FUNCTION_BLOCK "DRIVER_4C"   // FB249, SCL
TITLE = DRIVER_4C
{ S7_Optimized_Access := 'FALSE' }
AUTHOR : hugo
FAMILY : AUTOMAT
NAME : DRIVER4C
VERSION : 1.0
// driver_4C is a multi purpose driver.
// a rising edge on in switches from S0 state S1 and the next edge to state S2 and so on.
// in state S0 all outputs Q are FALSE.
// The stet of the Outputs in any state S? is configurable with setup variables.
// The variables S1..S5 define the states, while the sequence is terminated when a state Variable S? = 0.
// The lower bits 0..3 of the state vars S? are corresponding to the Outputs Q0..Q3
   VAR_INPUT
      IN : Bool;
      RST : Bool;
      Timeout : Time;
      SX : Array[1..7] of Byte;
   END_VAR
   VAR_OUTPUT
      SN : Int;
      Q0 : Bool;
      Q1 : Bool;
      Q2 : Bool;
      Q3 : Bool;
   END_VAR
   VAR
      off : TON;
      edge : Bool;
   END_VAR
   VAR_TEMP
      tSX : Byte;
      _SX AT tSX : Array[0..7] of Bool;
   END_VAR
   // SX[1] := B#16#01;
   // SX[2] := B#16#03;
   // SX[3] := B#16#07;
   // SX[4] := B#16#0F;
BEGIN


   IF #RST OR #off.Q THEN
       #SN := 0;
   ELSIF #IN AND NOT #edge THEN
       #SN := #SN + 1;
       IF #SN > 7 OR #SX[#SN] = 0 THEN #SN := 0; END_IF;
   END_IF;
   #edge := #IN;
   IF #SN > 0 THEN
       #tSX := #SX[#SN];  //so und nicht anders
       #Q0 := #_SX[0];
       #Q1 := #_SX[1];
       #Q2 := #_SX[2];
       #Q3 := #_SX[3];
   ELSE
       #Q0 := FALSE;
       #Q1 := FALSE;
       #Q2 := FALSE;
       #Q3 := FALSE;
   END_IF;

   (* maximaum timeout *)
   IF #Timeout > t#0s THEN #off(IN := #SN > 0, PT := #Timeout); END_IF;


   (* revision history
   hm  23. mar. 2009   rev 1.0
       original version

   *)
END_FUNCTION_BLOCK

FUNCTION "T_PLC_MS" : DWord   // FC64, SCL
TITLE = T_PLC_MS
{ S7_Optimized_Access := 'FALSE' }
AUTHOR : hugo
FAMILY : MEASURE
NAME : T_PLC_MS
VERSION : 1.2
// T_PLC_MS reads the internal PLC timer and return the time, it has the advantage to be able to set a debug mode 
// and speed up the counter to test the plc timer overrun which occurs every 50 days respectively 25 days at siemens S7
// this routine also allows to correct the behavior of s7 where the internal plc counter will not count all 32 bits.
// 
// uses: STIME [FB64],IDB_STIME [DB64]
BEGIN


   "IDB_STIME"(); 
   #T_PLC_MS := "IDB_STIME".tx; 
   (* hier muss die korrektur für step7 stattfinden
   plctime muss den vollen wertebereich von time ausnutzen:
   wenn bei step7 time -24tage bis plus 24 tage ist dann muss der timer auch beim überlauf auf -24tage springen 
   und auf keinen fall auf 0 !!!!
   für siemens muss ein weiterer fb im main eingebunden werden der sicherstellt das alle 32 bits durchgezählt werden.
   es kann nur ein fb sein den er muss sich das oberste (32te) bit merken.
   oder etwa spring s7 bei überlauf auf -24 tage????? dann wäre keine korrektur nötig.
   *)
   IF "debug" THEN
       #T_PLC_MS := DINT_TO_DWORD((DWORD_TO_DINT(SHL(IN:=#T_PLC_MS,N:="N") OR SHL(IN:=DWORD#1,N:="N"))-1) + DWORD_TO_DINT("offset_1"));
   END_IF;


   (* revision history
   hm  14.9.2007   rev 1.0
       original version

   hm  12. nov 2007    rev 1.1
       added temporaray variable tx because some compilers could not handle time() as an argument

   hm  16. nov. 2008   rev 1.2
       initialized constants with 0 for compatibility reasons
   *)
END_FUNCTION

FUNCTION "T_PLC_US" : DWord   // FC65, SCL
TITLE = T_PLC_US
{ S7_Optimized_Access := 'FALSE' }
AUTHOR : hugo
FAMILY : MEASURE
NAME : T_PLC_US
VERSION : 1.2
// T_PLC_US reads the internal PLC timer and return the time, it has the advantage to be able to set a debug mode 
// and speed up the counter to test the plc timer overrun which occurs every 50 days respectively 25 days at siemens S7
// this routine also allows to correct the behavior of s7 where the internal plc counter will not count all 32 bits.
// 
// uses: STIME [FB64],IDB_STIME [DB64]
BEGIN


   "IDB_STIME"(); 
   #T_PLC_US := DINT_TO_DWORD(DWORD_TO_DINT("IDB_STIME".tx) * 1000); 
   (* hier muss die korrektur für step7 stattfinden
   plctime muss den vollen wertebereich von time ausnutzen:
   wenn bei step7 time -24tage bis plus 24 tage ist dann muss der timer auch beim überlauf auf -24tage springen 
   und auf keinen fall auf 0 !!!!
   für siemens muss ein weiterer fb im main eingebunden werden der sicherstellt das alle 32 bits durchgezählt werden.
   es kann nur ein fb sein den er muss sich das oberste (32te) bit merken.
   oder etwa spring s7 bei überlauf auf -24 tage????? dann wäre keine korrektur nötig.
   *)
   IF "debug" THEN
       #T_PLC_US := DINT_TO_DWORD((DWORD_TO_DINT(SHL(IN:=#T_PLC_US,N:="N") OR SHL(IN:=DWORD#1,N:="N"))-1) + DWORD_TO_DINT("offset_1"));
   END_IF;


   (* revision history
   hm  14.9.2007   rev 1.0
       original version

   hm  12. nov 2007    rev 1.1
       added temporaray variable tx because some compilers could not handle time() as an argument

   hm  16. nov. 2008   rev 1.2
       initialized constants with 0 for compatibility reasons

   *)
END_FUNCTION

FUNCTION "INC" : Int   // FC90, SCL
TITLE = INC
{ S7_Optimized_Access := 'FALSE' }
AUTHOR : hugo
FAMILY : MATH
NAME : INC
VERSION : 1.1
// This is a increment function which increments the input X by the value D and compares the result with M.
// if the output exceeds M it will continue to count from 0 again.
   VAR_INPUT
      X : Int;
      D : Int;
      "M" : Int;
   END_VAR
BEGIN


     #INC := (#X + #D + #"M" + 1) MOD (#"M" + 1);

   (* revision history
   hm  7. feb 2007   REV 1.0
     original version

   hm  15. jan 2008  rev 1.1
     allow for neagtive increment

   *)
END_FUNCTION

FUNCTION "MULTIME" : Time   // FC203, SCL
TITLE = MULTIME
{ S7_Optimized_Access := 'FALSE' }
AUTHOR : hugo
FAMILY : TIDT
NAME : MULTIME
VERSION : 1.1
// multiplies a time by a real number and returns a time
   VAR_INPUT
      t : Time;
      "M" : Real;
   END_VAR
BEGIN


     #MULTIME := T_CONV(REAL_TO_DINT(DINT_TO_REAL(T_CONV(#t))*#"M"));

   (* revision history
   hm      2. oct 2006 rev 1.0
       original version

   hm      14. mar 2008    rev 1.1
       rounded the result after the last digit

   *)
END_FUNCTION

FUNCTION "MANUAL" : Bool   // FC409, SCL
TITLE = MANUAL
{ S7_Optimized_Access := 'FALSE' }
AUTHOR : hugo
FAMILY : AUTOMAT
NAME : MANUAL
VERSION : 1.0
// MANUAL is a manual override for digital signals.
// when on and off = FALSE, the output follows IN.
// ON = TRUE forces the output high, and OFF = TRUE forces the output low.
   VAR_INPUT
      IN : Bool;
      ON : Bool;
      OFF : Bool;
   END_VAR
BEGIN


   #MANUAL := NOT #OFF AND (#IN OR #ON);


   (* revision history
   hm  21. nov 2008    rev 1.0
       original version


   *)
END_FUNCTION

// ===== PLC "Engineering control"  Unspecific CPU S7 300 =====

VAR_GLOBAL CONSTANT   // PLC tag table "STEP7 classic symbols"
   "debug" : Bool := FALSE;
   "N" : Int := 0;
   "offset" : Int := 0;
   "offset_1" : DWord := 0;
END_VAR

TYPE "REAL2"
VERSION : 0.0
   STRUCT
      R1 : Real;
      RX : Real;
   END_STRUCT;
END_TYPE

DATA_BLOCK "IDB_STIME"   // DB64
{ S7_Optimized_Access := 'FALSE' }
AUTHOR : dalbi
FAMILY : MEASURE
VERSION : 0.0
// stored: InstanceOfName STIME
"STIME"
BEGIN
END_DATA_BLOCK

FUNCTION_BLOCK "CLK_PRG"   // FB52, SCL
TITLE = CLK_PRG
{ S7_Optimized_Access := 'FALSE' }
AUTHOR : hugo
FAMILY : GENERAT
NAME : CLK_PRG
VERSION : 1.3
// clk_prg uses the internal sps time to generate a clock with programmable period time.
// the period time is defined for 10ms .. 65s
// the first cycle after start is a clk pulse and then depending on the programmed period time a delay.
// every pulse is only valid for one cycle.
// the accuracy of clk_prg is depending on the accuracy of the system clock.
// 
// uses: T_PLC_MS [FC64]
//       STIME [FB64],IDB_STIME [DB64]
   VAR_INPUT
      PT : Time := T#10MS;
   END_VAR
   VAR_OUTPUT
      Q : Bool;
   END_VAR
   VAR
      init : Bool;
      last : Time;
      tx : Time;
   END_VAR
   VAR_TEMP
      TOP_SI : Struct
         EV_CLASS : Byte;
         EV_NUM : Byte;
         PRIORITY : Byte;
         NUM : Byte;
         TYP2_3 : Byte;
         TYP1 : Byte;
         ZI1 : Word;
         ZI2_3 : DWord;
      END_STRUCT;
      START_UP_SI : Struct
         EV_CLASS : Byte;
         EV_NUM : Byte;
         PRIORITY : Byte;
         NUM : Byte;
         TYP2_3 : Byte;
         TYP1 : Byte;
         ZI1 : Word;
         ZI2_3 : DWord;
      END_STRUCT;
      ERR : Int;
   END_VAR
BEGIN


   (* read actual startup info *)
   (* OB1_SCAN_1  BYTE  -  B#16#01: Abschluss des Neustarts (Warmstarts)
                        -  B#16#02: Abschluss des Wiederanlaufs
                        -  B#16#03: Abschluss des freien Zyklus
                        -  B#16#04: Abschluss des Kaltstarts
                        -  B#16#05: Erster OB 1-Zyklus der neuen Master-CPU nach 
                                    Master-Reserve-Umschaltung und STOP des 
                                    bisherigen Masters *)

   #ERR := RD_SINFO (TOP_SI => #TOP_SI, START_UP_SI => #START_UP_SI);

   (* read system time *)
   #tx := T_CONV(DWORD_TO_DINT("T_PLC_MS"()));

   (* reset last_time on system startup *)
   IF #TOP_SI.EV_NUM = 1 OR #TOP_SI.EV_NUM = 2 OR #TOP_SI.EV_NUM = 4 THEN 
       #init := false;
   END_IF;

   (* initialize on startup *)
   IF NOT #init THEN
       #init := TRUE;
       #last := #tx - #PT;
   END_IF;

   (* generate output pulse when next_pulse is reached *)
   #Q := #tx - #last >= #PT;
   IF #Q THEN #last := #tx; END_IF;


   (* revision hiostory

   hm 25 feb 2007  rev 1.1
       rewritten code for higher performance
       pt can now be changed during runtime

   hm  17. sep 2007    rev 1.2
       replaced time() with t_plc_ms() for compatibility reasons

   hm  25. oct. 2008   rev 1.3
       optimized code

   *)
END_FUNCTION_BLOCK

FUNCTION_BLOCK "STIME"   // FB64, SCL
TITLE = STIME
{ S7_Optimized_Access := 'FALSE' }
AUTHOR : dalbi
FAMILY : MEASURE
NAME : STIME
VERSION : 1.4
// this function block makes sure that the timer of a siemens sps counts from 0 - 2^32-1.
   VAR_OUTPUT
      tx : DWord;
      at_tx AT tx : Array[0..31] of Bool;
   END_VAR
   VAR
      last_time : DWord;
      bit31 : Bool;
      init : Bool := TRUE;
   END_VAR
   VAR_TEMP
      TOP_SI : Struct
         EV_CLASS : Byte;
         EV_NUM : Byte;
         PRIORITY : Byte;
         NUM : Byte;
         TYP2_3 : Byte;
         TYP1 : Byte;
         ZI1 : Word;
         ZI2_3 : DWord;
      END_STRUCT;
      START_UP_SI : Struct
         EV_CLASS : Byte;
         EV_NUM : Byte;
         PRIORITY : Byte;
         NUM : Byte;
         TYP2_3 : Byte;
         TYP1 : Byte;
         ZI1 : Word;
         ZI2_3 : DWord;
      END_STRUCT;
      ERR : Int;
   END_VAR
BEGIN


   (* this FB is only necessary for siemens sps
   the siemens sps timer counts from 0 to 2^31-1 and starts at 0 sfter overrun.
   this means that the bit 31 (the highest bit ) will never be used and therefore
   a problem arises when t2 - t1 is checked.
   t2 - t1 is always valid also in an timer overrun situation where the time t1 is very high and t2 is very low.
   the result of the subtraction t2 - t1 however is still valid.
   this calculation does not work for soiemens because the highest bit is not used.

   this module stores the highest bit, changes the highest bit at every overrun occurence and stuffs ther highest bit in the output.
   the output is then used by t_plc_us and t_plc_ms.

   the correction needs and fb and not a function because the value of the highest bit has to be stored.

   do never use this function block in a codesys environment. the timer in codesys is correct and runs from 0 to 2^32-1
   *)

   (* read actual startup info *)
   (* OB1_SCAN_1  BYTE  -  B#16#01: Abschluss des Neustarts (Warmstarts)
                        -  B#16#02: Abschluss des Wiederanlaufs
                        -  B#16#03: Abschluss des freien Zyklus
                        -  B#16#04: Abschluss des Kaltstarts
                        -  B#16#05: Erster OB 1-Zyklus der neuen Master-CPU nach 
                                    Master-Reserve-Umschaltung und STOP des 
                                    bisherigen Masters *)

   #ERR := RD_SINFO (TOP_SI => #TOP_SI, START_UP_SI => #START_UP_SI);

   (* reset last_time on system startup *)
   IF #TOP_SI.EV_NUM = 1 OR #TOP_SI.EV_NUM = 2 OR #TOP_SI.EV_NUM = 4 OR NOT #init THEN 
       #last_time := 0;
       #bit31 := false;
       #init := true;
   END_IF;

   (* read the system timer *)
   #tx := DINT_TO_DWORD(T_CONV(TIME_TCK()));

   (* check for overrun *)
   IF DWORD_TO_DINT(#tx) < DWORD_TO_DINT(#last_time) THEN
       (* an overrun has occured, change the value of the highest bit *)
       #bit31 := NOT #bit31;
   END_IF;

   (* stuff the highest bit into the timer value *)
   #at_tx[7] := #bit31;

   (* remember the last system time for the next overrun check *)
   #last_time := #tx;


   (* revision history
   DA  14.9.2007 rev 1.0
     original version

   DA  24.2.2008 rev 1.1
     added self reset on system startup

   DA   2.5.2008 rev 1.2
     corect a problem running under OB35

   DA  12.3.2009 rev 1.3
     corect a problem run on different CPUs

   DA  22.12.2009 rev 1.4
     corect a problem on startup
   *)
END_FUNCTION_BLOCK

FUNCTION_BLOCK "TP_X"   // FB69, SCL
TITLE = TP_X
{ S7_Optimized_Access := 'FALSE' }
AUTHOR : hugo
FAMILY : GENERAT
NAME : TP_R
VERSION : 1.3
// retriggerable edge triggered pulse similar to TP but with a retrigger function
// if the pt input is 0 then output is always low.
// 
// uses: T_PLC_MS [FC64]
//       STIME [FB64],IDB_STIME [DB64]
   VAR_INPUT
      IN : Bool;
      PT : Time;
   END_VAR
   VAR_OUTPUT
      Q : Bool;
      ET : Time;
   END_VAR
   VAR
      edge : Bool;
      start : Time;
      tx : Time;
   END_VAR
   VAR_TEMP
      TOP_SI : Struct
         EV_CLASS : Byte;
         EV_NUM : Byte;
         PRIORITY : Byte;
         NUM : Byte;
         TYP2_3 : Byte;
         TYP1 : Byte;
         ZI1 : Word;
         ZI2_3 : DWord;
      END_STRUCT;
      START_UP_SI : Struct
         EV_CLASS : Byte;
         EV_NUM : Byte;
         PRIORITY : Byte;
         NUM : Byte;
         TYP2_3 : Byte;
         TYP1 : Byte;
         ZI1 : Word;
         ZI2_3 : DWord;
      END_STRUCT;
      ERR : Int;
   END_VAR
BEGIN


   (* read actual startup info *)
   (* OB1_SCAN_1  BYTE  -  B#16#01: Abschluss des Neustarts (Warmstarts)
                        -  B#16#02: Abschluss des Wiederanlaufs
                        -  B#16#03: Abschluss des freien Zyklus
                        -  B#16#04: Abschluss des Kaltstarts
                        -  B#16#05: Erster OB 1-Zyklus der neuen Master-CPU nach 
                                    Master-Reserve-Umschaltung und STOP des 
                                    bisherigen Masters *)

   #ERR := RD_SINFO (TOP_SI => #TOP_SI, START_UP_SI => #START_UP_SI);

   (* read system_time *)
   #tx := T_CONV(DWORD_TO_DINT("T_PLC_MS"()));

   (* reset last_time on system startup *)
   IF #TOP_SI.EV_NUM = 1 OR #TOP_SI.EV_NUM = 2 OR #TOP_SI.EV_NUM = 4 THEN 
       #start := #tx;
   END_IF;

   (* rising edge trigger *)
   IF #IN AND NOT #edge THEN
       #start := #tx;
       #Q := #PT > t#0ms;
   ELSIF #Q THEN
       #ET := #tx - #start;
       IF #ET >= #PT THEN
           #Q := FALSE;
           #ET := t#0ms;
       END_IF;
   END_IF;
   #edge := #IN;


   (* revision history
   hm  4. aug 2006     rev 1.0
       original version

   hm  17. sep 2007    rev 1.1
       replaced time() with T_PLC_MS() for compatibility reasons

   hm  19. oct. 2008   rev 1.2
       renamed to TP_R to TP_X for compatibility reasons

   hm  17. dec. 2008   rev 1.3
       code optimized

   *)
END_FUNCTION_BLOCK

FUNCTION_BLOCK "PWM_DC"   // FB102, SCL
TITLE = PWM_DC
{ S7_Optimized_Access := 'FALSE' }
AUTHOR : oscat
FAMILY : SIGGEN
NAME : PWM_DC
VERSION : 1.4
// this signal generator generates a square wave signal which is specified by the frequency and the duty cycle
// 
// uses: CLK_PRG [FB52]
//       T_PLC_MS [FC64] 
//       STIME [FB64],IDB_STIME [DB64] 
//       TP_X [FB69]
   VAR_INPUT
      F : Real;
      DC : Real;
   END_VAR
   VAR_OUTPUT
      Q : Bool;
   END_VAR
   VAR
      clk : "CLK_PRG";
      pulse : "TP_X";
   END_VAR
   VAR_TEMP
      tmp : Real;
   END_VAR
BEGIN


   IF #F > 0.0 THEN
       #tmp := 1000.0 / #F;
       #clk(PT := T_CONV(REAL_TO_DINT(#tmp)));
       #pulse(IN := #clk.Q, PT := T_CONV(REAL_TO_DINT(#tmp * #DC)));

       #Q := #pulse.Q;
   END_IF;


   (* revision history

   hm  25. feb 2007    rev 1.1
       recoded in st for better performance and better portability

   hm  27. nov 2007    rev 1.2
       avoid divide by 0 when F = 0

   hm  19. oct. 2008   rev 1.3
       changed type TP_R to TP_X because of name change
       improved performance

   hm  11. mar. 2009   rev 1.4
       changed real constants to use dot syntax

   *)
END_FUNCTION_BLOCK

FUNCTION_BLOCK "CONTROL_SET1"   // FB142, SCL
TITLE = CONTROL_SET1
{ S7_Optimized_Access := 'FALSE' }
AUTHOR : hugo
FAMILY : CTRL
NAME : C_SET_1
VERSION : 1.1
// takahashi calculates controller parameters for P, PI and PID controllers based on the ziegler nichols method.
   VAR_INPUT
      Kt : Real;
      Tt : Real;
      PI : Bool;
      PID : Bool;
      P_K : Real := 5.0e-1;
      PI_K : Real := 4.5e-1;
      PI_TN : Real := 8.3e-1;
      PID_K : Real := 6.0e-1;
      PID_TN : Real := 5.0e-1;
      PID_TV : Real := 1.25e-1;
   END_VAR
   VAR_OUTPUT
      KP : Real;
      TN : Real;
      TV : Real;
      KI : Real;
      KD : Real;
   END_VAR
BEGIN


   IF #PI AND #PID THEN
       #KP := 0.0;
       #TN := 0.0;
       #TV := 0.0;
   ELSIF #PID THEN
       #KP := #PID_K * #Kt;
       #TN := #PID_TN * #Tt;
       #TV := #PID_TV * #Tt;
   ELSIF #PI THEN
       #KP := #PI_K * #Kt;
       #TN := #PI_TN * #Tt;
   ELSE
       #KP := #P_K * #Kt;
   END_IF;

   (* KI and KD are calculated *)
   IF #TN > 0.0 THEN #KI := #KP / #TN; ELSE #KI := 0.0; END_IF;
   #KD := #KP * #TV;


   (* revision history
   hm  4. nov 2007 rev 1.0
       original version

   hm  11. mar. 2009   rev 1.1
       real constants updated to new systax using dot

   *)
END_FUNCTION_BLOCK

FUNCTION_BLOCK "CONTROL_SET2"   // FB143, SCL
TITLE = CONTROL_SET2
{ S7_Optimized_Access := 'FALSE' }
AUTHOR : hugo
FAMILY : CTRL
NAME : C_SET_2
VERSION : 1.1
// takahashi calculates controller parameters for P, PI and PID controllers based on the ziegler nichols method.
   VAR_INPUT
      KS : Real;
      TU : Real;
      TG : Real;
      PI : Bool;
      PID : Bool;
      P_K : Real := 1.0e+0;
      PI_K : Real := 9.0e-1;
      PI_TN : Real := 3.33e+0;
      PID_K : Real := 1.2e+0;
      PID_TN : Real := 2.0e+0;
      PID_TV : Real := 5.0e-1;
   END_VAR
   VAR_OUTPUT
      KP : Real;
      TN : Real;
      TV : Real;
      KI : Real;
      KD : Real;
   END_VAR
   VAR
      TX : Real;
   END_VAR
BEGIN


   IF #TU > 0.0 AND #KS > 0.0 THEN #TX := #TG / #TU / #KS; END_IF;
   IF #PI AND #PID THEN
       #KP := 0.0;
       #TN := 0.0;
       #TV := 0.0;
   ELSIF #PID THEN
       #KP := #PID_K * #TX;
       #TN := #PID_TN * #TU;
       #TV := #PID_TV * #TU;
   ELSIF #PI THEN
       #KP := #PI_K * #TX;
       #TN := #PI_TN * #TU;
   ELSE
       #KP := #P_K * #TX;
   END_IF;

   (* KI and KD are calculated *)
   IF #TN > 0.0 THEN #KI := #KP / #TN; ELSE #KI := 0.0; END_IF;
   #KD := #KP * #TV;


   (* revision history
   hm  4. nov 2007 rev 1.0
       original version

   hm  11. mar. 2009   rev 1.1
       real constants updated to new systax using dot

   *)
END_FUNCTION_BLOCK

FUNCTION_BLOCK "CTRL_OUT"   // FB144, SCL
TITLE = CTRL_OUT
{ S7_Optimized_Access := 'FALSE' }
AUTHOR : hugo
FAMILY : CTRL
NAME : CTRL_OUT
VERSION : 1.1
   VAR_INPUT
      CI : Real;
      OFFSET : Real;
      MAN_IN : Real;
      LIM_L : Real;
      LIM_H : Real;
      MANUAL : Bool;
   END_VAR
   VAR_OUTPUT
      Y : Real;
      LIM : Bool;
   END_VAR
BEGIN


   #Y := SEL(G:=#MANUAL, IN0:=#CI, IN1:=#MAN_IN) + #OFFSET;

   (* Limit the output *)
   IF #Y > #LIM_L AND #Y < #LIM_H THEN
       #LIM := FALSE;
   ELSE
       #Y := LIMIT(MN:=#LIM_L, IN:=#Y, MX:=#LIM_H);
       #LIM := TRUE;
   END_IF;


   (* revision history
   hm  2. jun. 2008    rev 1.0
       original version

   hm  5. nov. 2008    rev 1.1
       optimized code
   *)
END_FUNCTION_BLOCK

FUNCTION_BLOCK "CTRL_PI"   // FB145, SCL
TITLE = CTRL_PI
{ S7_Optimized_Access := 'FALSE' }
AUTHOR : hugo
FAMILY : CTRL
NAME : CTRL_PI
VERSION : 2.0
// FT_PI is a PI controller with manual functionality.
// The PID controller works according to the fomula Y = e *(KP+ KI * INTEG(e) ) + offset, while e = set_point - actual.
// a rst will reset all internal data, while a switch to manual will cause the controller to follow the function Y = manual_in + offset.
// limit_h and Limit_l set the possible output range of Y.
// the output flags lim will signal that the output limits are active and overflow will signal that the integrator has reached its limits.
// 
// since rev 1.1 the "trapezregel is used for more accuracy.
// rev 1.2 added selective integratin which means the integrative component is only active within a small range of the target value 
// this avoids the integrator to go to limits while an input setpoint change happened and is only causing overshoots.
// the int_band is by default 100 which means the int is active all the time and if set to for example to 0.1 the integrator is only active
// while the input is between 0.9 and 1.1 of the set_point value.
// 
// default values for KP = 1, TN = 1, TV = 1, LIMIT_L = -1000, LIMIT_H = +1000.
// 
// uses: CTRL_IN [FC363]
//       DEAD_ZONE [FC365] 
//       FT_PIWL [FB161]
//       T_PLC_US [FC65] 
//       STIME [FB64],IDB_STIME [DB64] 
//       CTRL_OUT [FB144]
   VAR_INPUT
      ACT : Real;
      SET : Real;
      SUP : Real;
      OFS : Real;
      M_I : Real;
      MAN : Bool;
      RST : Bool;
      KP : Real := 1.0e+0;
      KI : Real := 1.0e+0;
      LL : Real := -1.0e+3;
      LH : Real := 1.0e+3;
   END_VAR
   VAR_OUTPUT
      Y : Real;
      DIFF : Real;
      LIM : Bool;
   END_VAR
   VAR
      pi : "FT_PIWL";
      co : "CTRL_OUT";
   END_VAR
BEGIN


   #DIFF := "CTRL_IN"(SET_POINT:=#SET, ACTUAL:=#ACT, NOISE:=#SUP);
   #pi(IN := #DIFF, KP := #KP, KI := #KI, LIM_L := #LL, LIM_H := #LH, RST := #RST);
   #co(CI := #pi.Y, OFFSET := #OFS, MAN_IN := #M_I, LIM_L := #LL, LIM_H := #LH, MANUAL := #MAN);
   #Y := #co.Y;
   #LIM := #co.LIM;


   (* revision history
   hm  31.10.2007      rev 1.0
       original version

   hm  3.11.2007       rev 1.1
       added noise input to filter noise
       added output diff
       set limit output false when output is within limits
       overfolw was not set correctly

   hm  5. jan 2008     rev 1.2
       improved performance

   hm  20. jun. 2008   rev 2.0
       rewritten using new modular approach

   *)
END_FUNCTION_BLOCK

FUNCTION_BLOCK "CTRL_PID"   // FB146, SCL
TITLE = CTRL_PID
{ S7_Optimized_Access := 'FALSE' }
AUTHOR : hugo
FAMILY : CTRL
NAME : CTRL_PID
VERSION : 2.0
// FT_PI is a PI controller with manual functionality.
// The PID controller works according to the fomula Y = e *(KP+ KI * INTEG(e) ) + offset, while e = set_point - actual.
// a rst will reset all internal data, while a switch to manual will cause the controller to follow the function Y = manual_in + offset.
// limit_h and Limit_l set the possible output range of Y.
// the output flags lim will signal that the output limits are active.
// 
// uses: CTRL_IN [FC363]
//       DEAD_ZONE [FC365] 
//       FT_PIDWL [FB159]
//       FT_PIWL [FB161] 
//       T_PLC_US [FC65]
//       STIME [FB64],IDB_STIME [DB64]
//       FT_DERIV [FB150] 
//       CTRL_OUT [FB144]
   VAR_INPUT
      ACT : Real;
      SET : Real;
      SUP : Real;
      OFS : Real;
      M_I : Real;
      MAN : Bool;
      RST : Bool;
      KP : Real := 1.0e+0;
      TN : Real := 1.0e+0;
      TV : Real := 1.0e+0;
      LL : Real := -1.0e+3;
      LH : Real := 1.0e+3;
   END_VAR
   VAR_OUTPUT
      Y : Real;
      DIFF : Real;
      LIM : Bool;
   END_VAR
   VAR
      pid : "FT_PIDWL";
      co : "CTRL_OUT";
   END_VAR
BEGIN


   #DIFF := "CTRL_IN"(SET_POINT:=#SET, ACTUAL:=#ACT, NOISE:=#SUP);
   #pid(IN := #DIFF, KP := #KP, TN := #TN, TV := #TV, LIM_L := #LL, LIM_H := #LH, RST := #RST);
   #co(CI := #pid.Y, OFFSET := #OFS, MAN_IN := #M_I, LIM_L := #LL, LIM_H := #LH, MANUAL := #MAN);
   #Y := #co.Y;
   #LIM := #co.LIM;



   (* revision history

   hm 1.12.2006        rev 1.1
       changed algorithm to trapezregel for higher accuracy.

   hm 3.1.2007     rev 1.2
       added integ_band to select when the integrator is active.

   hm  3.3.2007        rev 1.3
       added default values to inputs KP, TN, TV, LIMIT_L und LIMIT_H.

   hm 31.oct 2007  rev 1.4
       total rewrite of the module to avoid failures when one of the limits is 0

   hm  3.11.2007   rev 1.5
       added noise input to filter noise
       added output diff
       set limit output false when output is within limits
       overfolw was not set correctly

   hm  5. jan 2008 rev 1.6
       improved code for better performance
   *)
END_FUNCTION_BLOCK

FUNCTION_BLOCK "CTRL_PWM"   // FB147, SCL
TITLE = CTRL_PWM
{ S7_Optimized_Access := 'FALSE' }
AUTHOR : hugo
FAMILY : CTRL
NAME : CTRL_PWM
VERSION : 1.1
// uses: PWM_DC [FB102]
//       CLK_PRG [FB52] 
//       T_PLC_MS [FC64]
//       STIME [FB64],IDB_STIME [DB64]
//       TP_X [FB69]
   VAR_INPUT
      CI : Real;
      MAN_IN : Real;
      MANUAL : Bool;
      F : Real;
   END_VAR
   VAR_OUTPUT
      Q : Bool;
   END_VAR
   VAR
      PW : "PWM_DC";
   END_VAR
BEGIN


   #PW(F := #F, DC := SEL(G:=#MANUAL,IN0:=#CI,IN1:=#MAN_IN));
   #Q := #PW.Q;


   (* revision history
   hm  3. jun. 2008    rev 1.0
       original version

   hm  21. oct. 2008    rev 1.1
       optimized code
   *)
END_FUNCTION_BLOCK

FUNCTION_BLOCK "DEAD_BAND_A"   // FB148, SCL
TITLE = DEAD_BAND_A
{ S7_Optimized_Access := 'FALSE' }
AUTHOR : hugo
FAMILY : CTRL
NAME : DEADBD_A
VERSION : 1.1
// DEAD_BAND ist eine lineare Übertragungsfunktion mit Totzone. Die Funktion verschiebt den positiven Teil der Kurve um -L und den negativen Teil der Kurve um +L.
// DEAD_BAND = X wenn Abs(X) > L wenn Abs(X) > L
// DEAD_BAND = 0 wenn Abs(X) <= L
// Die Breite der Totzone wird automatisch aus dem Signalrauschen errechnet.
// 
// uses: FT_PT1 [FB162]
//       T_PLC_US [FC65] 
//       STIME [FB64],IDB_STIME [DB64] 
//       MULTIME [FC203]
   VAR_INPUT
      X : Real;
      T : Time;
      KL : Real := 1.0e+0;
      LM : Real;
   END_VAR
   VAR_OUTPUT
      Y : Real;
      L : Real;
   END_VAR
   VAR
      tp1 : "FT_PT1";
      tp2 : "FT_PT1";
   END_VAR
BEGIN


   (* filter the input signal *)
   #tp1(in := #X, T:= #T);

   (* filter the HF portion to generate a stable L *)
   #tp2(in := ABS(#tp1.out - #X), T := "MULTIME"(t:=#T,M:=4.0));

   (* now we determine L which is half the width of the dead band *)
   #L := MIN(IN1:=#KL * #tp2.out,IN2:=#LM);

   IF #X > #L THEN
       #Y := #X - #L;
   ELSIF #X < -#L THEN
       #Y := #X + #L;
   ELSE
       #Y := 0.0;
   END_IF;


   (* revision history
   hm  14. jun. 2008   rev 1.0
       original version

   hm  11. mar. 2009   rev 1.1
       real constants updated to new systax using dot

   *)
END_FUNCTION_BLOCK

FUNCTION_BLOCK "DEAD_ZONE2"   // FB149, SCL
TITLE = DEAD_ZONE2
{ S7_Optimized_Access := 'FALSE' }
AUTHOR : hugo
FAMILY : CTRL
NAME : DEADZ2
VERSION : 1.1
// dead_zone2 is a linear transfer function which follows a linear function except for x is close to 0.
// Y = X if abs(x) > L.
// for values of 0 +/. L a hysteresis function will hold the output at + or - L.
   VAR_INPUT
      X : Real;
      L : Real;
   END_VAR
   VAR_OUTPUT
      Y : Real;
   END_VAR
BEGIN


   IF ABS(#X) > #L THEN
       #Y := #X;
   ELSIF #Y > 0.0 THEN
       #Y := #L;
   ELSE
       #Y := -#L;
   END_IF;


   (* revision history

   hm  12. feb. 2007   rev 1.0
       original version

   hm  11. mar. 2009   rev 1.1
       real constants updated to new systax using dot

   *)
END_FUNCTION_BLOCK

FUNCTION_BLOCK "FT_DERIV"   // FB150, SCL
TITLE = FT_DERIV
{ S7_Optimized_Access := 'FALSE' }
AUTHOR : hugo
FAMILY : CTRL
NAME : DERIV
VERSION : 1.5
// FT_deriv calculates the derivate over the signal "in" with Faktor "K".
// a run input enables or stops the calculation, if left unconnected its true and therfore the calculation is executed.
// if K is not specified the default is 1.
// 
// uses: T_PLC_US [FC65]
//       STIME [FB64],IDB_STIME [DB64]
   VAR_INPUT
      in : Real;
      K : Real := 1.0e+0;
      run : Bool := TRUE;
   END_VAR
   VAR_OUTPUT
      out : Real;
   END_VAR
   VAR
      old : Real;
      tx : DWord;
      last : DWord;
      init : Bool;
      tc : Real;
   END_VAR
   VAR_TEMP
      TOP_SI : Struct
         EV_CLASS : Byte;
         EV_NUM : Byte;
         PRIORITY : Byte;
         NUM : Byte;
         TYP2_3 : Byte;
         TYP1 : Byte;
         ZI1 : Word;
         ZI2_3 : DWord;
      END_STRUCT;
      START_UP_SI : Struct
         EV_CLASS : Byte;
         EV_NUM : Byte;
         PRIORITY : Byte;
         NUM : Byte;
         TYP2_3 : Byte;
         TYP1 : Byte;
         ZI1 : Word;
         ZI2_3 : DWord;
      END_STRUCT;
      ERR : Int;
   END_VAR
BEGIN


   (* read actual startup info *)
   (* OB1_SCAN_1  BYTE  -  B#16#01: Abschluss des Neustarts (Warmstarts)
                        -  B#16#02: Abschluss des Wiederanlaufs
                        -  B#16#03: Abschluss des freien Zyklus
                        -  B#16#04: Abschluss des Kaltstarts
                        -  B#16#05: Erster OB 1-Zyklus der neuen Master-CPU nach 
                                    Master-Reserve-Umschaltung und STOP des 
                                    bisherigen Masters *)

   #ERR := RD_SINFO (TOP_SI => #TOP_SI, START_UP_SI => #START_UP_SI);

   (* reset last_time on system startup *)
   IF #TOP_SI.EV_NUM = 1 OR #TOP_SI.EV_NUM = 2 OR #TOP_SI.EV_NUM = 4 THEN 
       #init := FALSE;
   END_IF;

   (* read system time *)
   #tx := "T_PLC_US"();
   #tc := DINT_TO_REAL(DWORD_TO_DINT(#tx) - DWORD_TO_DINT(#last));

   (* init on firsat startup *)
   IF NOT #init THEN
       #init := TRUE;
       #old := #in;
   ELSIF #run AND #tc > 0.0 THEN 
       #out := (#in - #old) / #tc * 1000000.0 * #K;
       #old := #in;
   ELSE
       #out := 0.0;
   END_IF;

   #last := #tx;


   (*
   hm 3.1.2007         rev 1.1
       added init code for startup
       set the default for K to 1

   hm  15. sep 2007    rev 1.2
       replaced Time() with T_PLC_US for compatibility and performance reasons
       increased accuracy and work in microseconds internally

   hm 29 oct 2007  rev 1.3
       prohibit calculation when tx - last = 0 to avoid division by 0 and increase accuracy on fast systems

   hm  6. nov. 2008    rev 1.4
       improved performance

   hm  11. mar. 2009   rev 1.5
       inproved code
   *)
END_FUNCTION_BLOCK

FUNCTION_BLOCK "FT_IMP"   // FB151, SCL
TITLE = FT_IMP
{ S7_Optimized_Access := 'FALSE' }
AUTHOR : hugo
FAMILY : CTRL
NAME : IMP
VERSION : 1.1
// FT_IMP is   an impulse filter (high pass filter) with the time T and factor K.
// 
// uses: FT_PT1 [FB162]
//       T_PLC_US [FC65] 
//       STIME [FB64],IDB_STIME [DB64]
   VAR_INPUT
      in : Real;
      T : Time;
      K : Real := 1.0e+0;
   END_VAR
   VAR_OUTPUT
      out : Real;
   END_VAR
   VAR
      t_1 : "FT_PT1";
   END_VAR
BEGIN


     #t_1(in:= #in, T:=#T);
     #out := (#in - #t_1.out) * #K;

   (*
   hm 3.1.2007  rev 1.1
     added factor K

   *)
END_FUNCTION_BLOCK

FUNCTION_BLOCK "FT_INT"   // FB152, SCL
TITLE = FT_INT
{ S7_Optimized_Access := 'FALSE' }
AUTHOR : hugo
FAMILY : CTRL
NAME : _INT
VERSION : 2.2
// FT_int is an integrator with input IN and factor K.
// integration is only done while run = true, if run is false integration is stopped and the out remains at the last value.
// if run is left unconnected, run is considered true by the function block.
// the output ET will display the total integration time from last reset.
// the out_min and out_max values can be set to ,imit the output value range. 
// the default for K is 1.
// 
// uses: INTEGRATE [FB237]
//       T_PLC_MS [FC64] 
//       STIME [FB64],IDB_STIME [DB64]
   VAR_INPUT
      IN : Real;
      K : Real := 1.0e+0;
      RUN : Bool := TRUE;
      RST : Bool;
      OUT_MIN : Real := -1.0e+37;
      OUT_MAX : Real := 1.0e+37;
   END_VAR
   VAR_OUTPUT
      OUT : Real;
      LIM : Bool;
   END_VAR
   VAR
      INTeg : "INTEGRATE";
   END_VAR
BEGIN


   IF #RST THEN
       #OUT := 0.0;
   ELSE
       #INTeg(X := #IN, E := #RUN, K := #K, Y := #OUT);
   END_IF;

   (* limit the outputs *)
   IF #OUT >= #OUT_MAX THEN
       #OUT := #OUT_MAX;
       #LIM := TRUE;
   ELSIF #OUT <= #OUT_MIN THEN
       #OUT := #OUT_MIN;
       #LIM := TRUE;
   ELSE
       #LIM := FALSE;
   END_IF;


   (*
   hm 13.12.2006   rev 1.1
       changed to "trapezregel" which increases accuracy
       before out := out + in * time new: out := out + (in + in_last) / 2 * time

   hm 15.1.2007        rev 1.2
       added default for k to be 1.

   hm  15.9.2007       rev 1.3
       replaced time() with T_PLC_US for compatibility and performance reason
       increased internal accuracy to microseconds

   hm 29. oct 2007     rev 1.4
       changed code so int will not be called is time difference is 0 to increase accuracy on systems
       with cycle times below 1ms

   hm  2. dec 2007     rev 1.5
       changed code for better performance

   hm  5. jan 2008     rev 1.6
       further improvements in performance

   hm  8. feb 2008     rev 1.7
       deleted limits +/- 1000 now limit is the range of real
       added variables out1 and out2 to extend the resolution
       corrected an error with elapsed time
       deleted unusfull output ET

   hm  13. mar 2008    rev 1.8
       changed preset value out_min to -1e37.
       stop integrator at the limits.

   hm  16. mar 2008    rev 1.9
       added type conversion to avoid warning under codesys 3.0

   hm  2. jun. 2008    rev 2.0
       rewritten with clear code
       limits can now be set without run

   hm  3. nov. 2008    rev 2.1
       optimized code using INTEGRATE and LIMX

   hm  10. mar. 2009   rev 2.2
       removed nested comments
   *)
END_FUNCTION_BLOCK

FUNCTION_BLOCK "FT_INT2"   // FB153, SCL
TITLE = FT_INT2
{ S7_Optimized_Access := 'FALSE' }
AUTHOR : hugo
FAMILY : CTRL
NAME : FT_INT2
VERSION : 1.2
// FT_int is an integrator with input IN and factor K.
// integration is only done while run = true, if run is false integration is stopped and the out remains at the last value.
// if run is left unconnected, run is considered true by the function block.
// the out_min and out_max values can be set to ,imit the output value range. 
// the default for K is 1.
// FT_INT2 has double presision accuracy (14 disgits).
// 
// uses: REAL2 [UDT11]
//       R2_SET [FC147]
//       INTEGRATE [FB237]
//       T_PLC_MS [FC64] 
//       STIME [FB64],IDB_STIME [DB64] 
//       R2_ADD [FC144]
   VAR_INPUT
      IN : Real;
      K : Real := 1.0e+0;
      RUN : Bool := TRUE;
      RST : Bool;
      OUT_MIN : Real := -1.0e+38;
      OUT_MAX : Real := 1.0e+38;
   END_VAR
   VAR_OUTPUT
      OUT : Real;
      LIM : Bool;
   END_VAR
   VAR
      integ : "INTEGRATE";
      ix : Real;
      val : "REAL2";
   END_VAR
BEGIN


   IF #RST THEN
       #val := "R2_SET"(0.0);
       #OUT := 0.0;
   ELSE
       #integ(X := #IN, E := #RUN, K := #K, Y := #ix);
       #val := "R2_ADD"(X:=#val, Y:=#ix);
       #ix := 0.0;
       #OUT := #val.RX;
   END_IF;

   (* check output for limits *)
   IF #OUT > #OUT_MIN AND #OUT < #OUT_MAX THEN
       #LIM := FALSE;
   ELSE
       #OUT := LIMIT(MN:=#OUT_MIN, IN:=#OUT, MX:=#OUT_MAX);
       #val := "R2_SET"(#OUT);
       #LIM := TRUE;
   END_IF;


   (*  revision history
   hm  2. jun. 2008    rev 1.0
       original version

   hm  5. nov. 2008    rev 1.1
       rewritten code using integrate

   hm  11. mar. 2009   rev 1.2
       real constants updated to new systax using dot

   *)
END_FUNCTION_BLOCK

FUNCTION_BLOCK "FT_PD"   // FB154, SCL
TITLE = FT_PD
{ S7_Optimized_Access := 'FALSE' }
AUTHOR : hugo
FAMILY : CTRL
NAME : FT_PD
VERSION : 1.0
// FT_PD is a PD controller.
// The PD controller works according to the fomula Y = KP *(IN + DERIV(e) ).
// 
// uses: FT_DERIV [FB150]
//       T_PLC_US [FC65] 
//       STIME [FB64],IDB_STIME [DB64]
   VAR_INPUT
      IN : Real;
      KP : Real := 1.0e+0;
      TV : Real := 1.0e+0;
   END_VAR
   VAR_OUTPUT
      Y : Real;
   END_VAR
   VAR
      diff : "FT_DERIV";
   END_VAR
BEGIN


   (* run differentiator *)
   #diff(in := #IN, K := #TV);

   (* combine both values *)
   #Y := #KP * (#diff.out + #IN);



   (* revision history
   hm  3. jun. 2008    rev 1.0
       original version


   *)
END_FUNCTION_BLOCK

FUNCTION_BLOCK "FT_PDT1"   // FB155, SCL
TITLE = FT_PDT1
{ S7_Optimized_Access := 'FALSE' }
AUTHOR : hugo
FAMILY : CTRL
NAME : FT_PDT1
VERSION : 1.0
// FT_PD is a PD controller.
// The PD controller works according to the fomula Y = KP *(IN + DERIV(e) ).
// 
// uses: FT_DERIV [FB150]
//       T_PLC_US [FC65] 
//       STIME [FB64],IDB_STIME [DB64] 
//       FT_PT1 [FB162]
   VAR_INPUT
      IN : Real;
      KP : Real := 1.0e+0;
      TV : Real := 1.0e+0;
      _T1 : Real := 1.0e+0;
   END_VAR
   VAR_OUTPUT
      Y : Real;
   END_VAR
   VAR
      diff : "FT_DERIV";
      TP : "FT_PT1";
   END_VAR
BEGIN


   (* run differentiator *)
   #diff(in := #IN, K := #TV);

   (* Run PT1 filter *)
   #TP(in := #diff.out, T := T_CONV(REAL_TO_DINT(#_T1)));

   (* combine both values *)
   #Y := #KP * (#TP.out + #IN);



   (* revision history
   hm  3. jun. 2008    rev 1.0
       original version


   *)
END_FUNCTION_BLOCK

FUNCTION_BLOCK "FT_PI"   // FB156, SCL
TITLE = FT_PI
{ S7_Optimized_Access := 'FALSE' }
AUTHOR : hugo
FAMILY : CTRL
NAME : PI
VERSION : 2.0
// FT_PI is a PI controller.
// The PID controller works according to the fomula Y = IN *(KP+ KI * INTEG(e) ).
// a rst will reset the integrator to 0
// ilim_h and iLim_l set the possible output range of the internal integrator.
// the output flags lim will signal that the output limits are active.
// 
// default values for KP = 1, KI = 1, ILIM_L = -1E37, iLIM_H = +1E38.
//  
// uses: FT_INT [FB152]
//       INTEGRATE [FB237] 
//       T_PLC_MS [FC64]
//       STIME [FB64],IDB_STIME [DB64]
   VAR_INPUT
      IN : Real;
      KP : Real := 1.0e+0;
      KI : Real := 1.0e+0;
      ILIM_L : Real := -1.0e+38;
      ILIM_H : Real := 1.0e+38;
      IEN : Bool := TRUE;
      RST : Bool;
   END_VAR
   VAR_OUTPUT
      Y : Real;
      LIM : Bool;
   END_VAR
   VAR
      integ : "FT_INT";
   END_VAR
BEGIN


   (* run integrator *)
   #integ(IN := #IN, K := #KI, RUN := #IEN, RST := #RST, OUT_MIN := #ILIM_L, OUT_MAX := #ILIM_H);
   (* check if integrator has reached its limits and set overflow *)
   #LIM := #integ.LIM;
   #Y := #KP * #IN + #integ.OUT;



   (* revision history
   hm  3. jun. 2008    rev 2.0
       original version


   *)
END_FUNCTION_BLOCK

FUNCTION_BLOCK "FT_PID"   // FB157, SCL
TITLE = FT_PID
{ S7_Optimized_Access := 'FALSE' }
AUTHOR : hugo
FAMILY : CTRL
NAME : PID
VERSION : 2.1
// FT_PI is a PI controller.
// The PID controller works according to the fomula Y = IN *(KP+ KI * INTEG(e) ).
// a rst will reset the integrator to 0
// ilim_h and iLim_l set the possible output range of the internal integrator.
// the output flags lim will signal that the output limits are active.
// 
// default values for KP = 1, KI = 1, ILIM_L = -1E37, iLIM_H = +1E38.
// 
// uses: FT_INT [FB152]
//       INTEGRATE [FB237] 
//       T_PLC_MS [FC64]
//       STIME [FB64],IDB_STIME [DB64]
//       FT_DERIV [FB150]
//       T_PLC_US [FC65]
   VAR_INPUT
      IN : Real;
      KP : Real := 1.0e+0;
      TN : Real := 1.0e+0;
      TV : Real := 1.0e+0;
      ILIM_L : Real := -1.0e+38;
      ILIM_H : Real := 1.0e+38;
      IEN : Bool := TRUE;
      RST : Bool;
   END_VAR
   VAR_OUTPUT
      Y : Real;
      LIM : Bool;
   END_VAR
   VAR
      integ : "FT_INT";
      diff : "FT_DERIV";
   END_VAR
BEGIN


   (* run integrator only if TN > 0 *)
   IF #TN > 0.0 THEN
       #integ(IN := #IN, K := 1.0 / #TN, RUN := #IEN, RST := #RST, OUT_MIN := #ILIM_L, OUT_MAX := #ILIM_H);
   ELSE
       #integ(RST := FALSE);
   END_IF;

   (* run differentiator *)
   #diff(in := #IN, K := #TV);

   (* combine both values *)
   #Y := #KP * (#integ.OUT + #diff.out + #IN);

   (* check if integrator has reached its limits and set overflow *)
   #LIM := #integ.LIM;


   (* revision history
   hm 3. jun. 2008     rev 2.0
       original version

   hm  11. mar. 2009   rev 2.1
       real constants updated to new systax using dot

   *)
END_FUNCTION_BLOCK

FUNCTION_BLOCK "FT_PIDW"   // FB158, SCL
TITLE = FT_PIDW
{ S7_Optimized_Access := 'FALSE' }
AUTHOR : hugo
FAMILY : CTRL
NAME : FT_PIDW
VERSION : 1.2
// FT_PIDW is a PID controller with dynamic wind_up reset.
// The PID controller works according to the fomula Y = KP *(IN + KI * INTEG(e) + DERIV(e) ).
// a rst will reset the integrator to 0
// lim_h and Lim_l set the possible output range of the internal integrator.
// the output flags lim will signal that the output limits are active.
// 
// default values for KP = 1, KI = 1, ILIM_L = -1E37, iLIM_H = +1E38.
// 
// uses: INTEGRATE [FB237]
//       T_PLC_MS [FC64] 
//       STIME [FB64],IDB_STIME [DB64] 
//       FT_DERIV [FB150]
//       T_PLC_US [FC65]
   VAR_INPUT
      IN : Real;
      KP : Real := 1.0e+0;
      TN : Real := 1.0e+0;
      TV : Real := 1.0e+0;
      LIM_L : Real := -1.0e+38;
      LIM_H : Real := 1.0e+38;
      RST : Bool;
   END_VAR
   VAR_OUTPUT
      Y : Real;
      LIM : Bool;
   END_VAR
   VAR
      integ : "INTEGRATE";
      diff : "FT_DERIV";
      YI : Real;
   END_VAR
BEGIN


   (* run the integrator *)
   IF #TN = 0.0 OR #RST THEN
       #integ(E := FALSE, Y := #YI);
       #YI := 0.0;
   ELSE
       #integ(X := #IN, K := 1.0 / #TN, E := NOT #LIM, Y := #YI);
   END_IF;

   (* add up integrator and linear part *)
   #Y := #KP * (#IN + #YI);

   (* run differentiator *)
   #diff(in := #IN, K := #TV);

   (* set lim before differentiator is added to stop integrator if necessary *)
   IF #Y > #LIM_L AND #Y < #LIM_H THEN
       #LIM := FALSE;
   ELSE
       #LIM := TRUE;
   END_IF;

   (* add differential part and limit output Y *)

   #Y := LIMIT(MN:=#LIM_L, IN:=#Y + #KP * #diff.out, MX:=#LIM_H);


   (* revision history
   hm 3. jun. 2008     rev 1.0
       original version

   hm  5. nov. 2008  rev 1.1
       changed code to use integrate

   hm  11. mar. 2009   rev 1.2
       real constants updated to new systax using dot

   *)
END_FUNCTION_BLOCK

FUNCTION_BLOCK "FT_PIDWL"   // FB159, SCL
TITLE = FT_PIDWL
{ S7_Optimized_Access := 'FALSE' }
AUTHOR : hugo
FAMILY : CTRL
NAME : FT_PIDWL
VERSION : 1.3
// FT_PIDW is a PID controller with dynamic wind_up reset.
// The PID controller works according to the fomula Y = KP *(IN + KI * INTEG(e) + DERIV(e) ).
// a rst will reset the integrator to 0
// lim_h and Lim_l set the possible output range of the internal integrator.
// the output flags lim will signal that the output limits are active.
// 
// default values for KP = 1, KI = 1, ILIM_L = -1E37, iLIM_H = +1E38.
// 
// uses: FT_PIWL [FB161]
//       T_PLC_US [FC65] 
//       STIME [FB64],IDB_STIME [DB64] 
//       FT_DERIV [FB150]
   VAR_INPUT
      IN : Real;
      KP : Real := 1.0e+0;
      TN : Real := 1.0e+0;
      TV : Real := 1.0e+0;
      LIM_L : Real := -1.0e+38;
      LIM_H : Real := 1.0e+38;
      RST : Bool;
   END_VAR
   VAR_OUTPUT
      Y : Real;
      LIM : Bool;
   END_VAR
   VAR
      piwl : "FT_PIWL";
      diff : "FT_DERIV";
   END_VAR
BEGIN


   (* if rst then *)
   IF #RST THEN
       #piwl(RST := TRUE);
       #piwl.RST := FALSE;
   ELSE
       (* run PIWL controller first *)
       (* we need to check if TN = 0 and do alternative calls *)
       IF #TN = 0.0 THEN
         #piwl(IN := #IN * #KP, KP := 1.0, KI := 0.0, LIM_L := #LIM_L, LIM_H := #LIM_H);
       ELSE
         #piwl(IN := #IN * #KP, KP := 1.0, KI := 1.0 / #TN, LIM_L := #LIM_L, LIM_H := #LIM_H);
       END_IF;

       (* run differentiator and add_to_output *)
       #diff(in := #IN, K := #KP * #TV);
       #Y := #piwl.Y + #diff.out;

       (* limit the output *)
       IF #Y < #LIM_L THEN
           #LIM := TRUE;
           #Y := #LIM_L;
       ELSIF #Y > #LIM_H THEN
           #LIM := TRUE;
           #Y := #LIM_H;
       ELSE
           #LIM := FALSE;
       END_IF;
   END_IF;


   (* revision history
   hm 13. jun. 2008  rev 1.0
     original version

   hm  25. jan 2008  rev 1.1
     multiply differential part with KP

   hm  11. mar. 2009 rev 1.2
     real constants updated to new systax using dot

   hm  13. nov. 2009 rev 1.3
     fixed code for negative KP

   *)
END_FUNCTION_BLOCK

FUNCTION_BLOCK "FT_PIW"   // FB160, SCL
TITLE = FT_PIW
{ S7_Optimized_Access := 'FALSE' }
AUTHOR : hugo
FAMILY : CTRL
NAME : FT_PIW
VERSION : 1.0
// FT_PIW is a PI controller.
// The PID controller works according to the fomula Y = IN *(KP+ KI * INTEG(e) ).
// a rst will reset the integrator to 0
// ilim_h and iLim_l set the possible output range of the internal integrator.
// the output flag lim will signal that the output limits are active.
// the controller is equipped with anti wind_up circuitry that stops the integrator when lim_h or lim_l is reached
// 
// default values for KP = 1, KI = 1, ILIM_L = -1E37, iLIM_H = +1E38.
// 
// uses: FT_INT [FB152]
//       INTEGRATE [FB237] 
//       T_PLC_MS [FC64]
//       STIME [FB64],IDB_STIME [DB64]
   VAR_INPUT
      IN : Real;
      KP : Real := 1.0e+0;
      KI : Real := 1.0e+0;
      LIM_L : Real := -1.0e+38;
      LIM_H : Real := 1.0e+38;
      RST : Bool;
   END_VAR
   VAR_OUTPUT
      Y : Real;
      LIM : Bool;
   END_VAR
   VAR
      integ : "FT_INT";
   END_VAR
BEGIN


   (* run integrator *)
   #integ(IN := #IN, K := #KI, RUN := NOT #LIM, RST := #RST);

   (* set output value *)
   #Y := #KP * #IN + #integ.OUT;

   (* check for limits and set integrator for anti wind up *)
   IF #Y < #LIM_L THEN
       #Y := #LIM_L;
       #LIM := TRUE;
   ELSIF #Y > #LIM_H THEN
       #Y := #LIM_H;
       #LIM := TRUE;
   ELSE
       #LIM := FALSE;
   END_IF;



   (* revision history
   hm  3. jun. 2008    rev 1.0
       original version


   *)
END_FUNCTION_BLOCK

FUNCTION_BLOCK "FT_PIWL"   // FB161, SCL
TITLE = FT_PIWL
{ S7_Optimized_Access := 'FALSE' }
AUTHOR : hugo
FAMILY : CTRL
NAME : FT_PIWL
VERSION : 1.3
// FT_PIWL is a PI controller.
// The PID controller works according to the fomula Y = IN *(KP+ KI * INTEG(e) ).
// a rst will reset the integrator to 0
// lim_h and Lim_l set the possible output range of the controller.
// the output flag lim will signal that the output limits are active.
// the integrator ist equipped with anti wind-up circuitry which limits trhe total output ranke to lim_l and lim_h
// 
// default values for KP = 1, KI = 1, ILIM_L = -1E37, iLIM_H = +1E38.
// 
// uses: T_PLC_US [FC65]
//       STIME [FB64],IDB_STIME [DB64]
   VAR_INPUT
      IN : Real;
      KP : Real := 1.0e+0;
      KI : Real := 1.0e+0;
      LIM_L : Real := -1.0e+38;
      LIM_H : Real := 1.0e+38;
      RST : Bool;
   END_VAR
   VAR_OUTPUT
      Y : Real;
      LIM : Bool;
   END_VAR
   VAR
      init : Bool;
      tx : DWord;
      tc : Real;
      t_last : DWord;
      in_last : Real;
      i : Real;
      p : Real;
   END_VAR
BEGIN


   (* initialize at power_up *)
   IF NOT #init OR #RST THEN
       #init := TRUE;
       #in_last := #IN;
       #t_last := "T_PLC_US"();
       #i := 0.0;
       #tc := 0.0;
   ELSE
       (* read last cycle time in Microseconds *)
       #tx := "T_PLC_US"();
       #tc := DINT_TO_REAL(DWORD_TO_DINT(#tx) - DWORD_TO_DINT(#t_last));
       #t_last := #tx;

       (* calculate proportional part *)
       #p := #KP * #IN;

       (* run integrator *)
       #i := (#IN + #in_last) * 5.0E-7 * #KI * #tc + #i;
       #in_last := #IN;

       (* calculate output Y *)
       #Y := #p + #i;

       (* check output for limits *)
       IF #Y >= #LIM_H THEN
           #Y := #LIM_H;
           IF #KI <> 0.0 THEN  
               #i := #LIM_H - #p; 
           ELSE
               #i := 0.0;
           END_IF;
           #LIM := TRUE;
       ELSIF #Y <= #LIM_L THEN
           #Y := #LIM_L;
           IF #KI <> 0.0 THEN 
               #i := #LIM_L - #p; 
           ELSE
               #i := 0.0;
           END_IF;
           #LIM := TRUE;
       ELSE
           #LIM := FALSE;
       END_IF;
   END_IF;


   (* revision history
   hm 13. jun. 2008    rev 1.0
       original version

   hm  27. oct. 2008   rev 1.1
       integrator will not be adjusted when ki = 0

   hm  25. jan 2009    rev 1.2
       module will also work with negative K

   hm  11. mar. 2009   rev 1.3
       real constants updated to new systax using dot

   *)
END_FUNCTION_BLOCK

FUNCTION_BLOCK "FT_PT1"   // FB162, SCL
TITLE = FT_PT1
{ S7_Optimized_Access := 'FALSE' }
AUTHOR : hugo
FAMILY : CTRL
NAME : PT1
VERSION : 1.11
// FT_PT1 is an low pass filter with a programmable time T and faktor K.
// 
// uses: T_PLC_US [FC65]
//       STIME [FB64],IDB_STIME [DB64]
   VAR_INPUT
      in : Real;
      T : Time;
      K : Real := 1.0e+0;
   END_VAR
   VAR_OUTPUT
      out : Real;
   END_VAR
   VAR
      last : DWord;
      tx : DWord;
      init : Bool;
   END_VAR
BEGIN


   (* read system time *)
   #tx := "T_PLC_US"();